REGION Network 92
   RUNG wire#powerrail
      Contact( "Carrier_14_Status.8" )
      Coil( "EMS".Carrier[14].SDC_IN.CrashDetectStatus )
   END_RUNG
   // the same network as SCL:
   "EMS".Carrier[14].SDC_IN.CrashDetectStatus := "Carrier_14_Status.8";
END_REGION

REGION Network 93
   RUNG wire#powerrail
      Contact( "Carrier_14_Status.9" )
      Coil( "EMS".Carrier[14].SDC_IN.EncoderCommFault )
   END_RUNG
   // the same network as SCL:
   "EMS".Carrier[14].SDC_IN.EncoderCommFault := "Carrier_14_Status.9";
END_REGION

REGION Network 94
   RUNG wire#powerrail
      Contact( "Carrier_14_Status.10" )
      Coil( "EMS".Carrier[14].SDC_IN.DriveCommFault )
   END_RUNG
   // the same network as SCL:
   "EMS".Carrier[14].SDC_IN.DriveCommFault := "Carrier_14_Status.10";
END_REGION

REGION Network 95
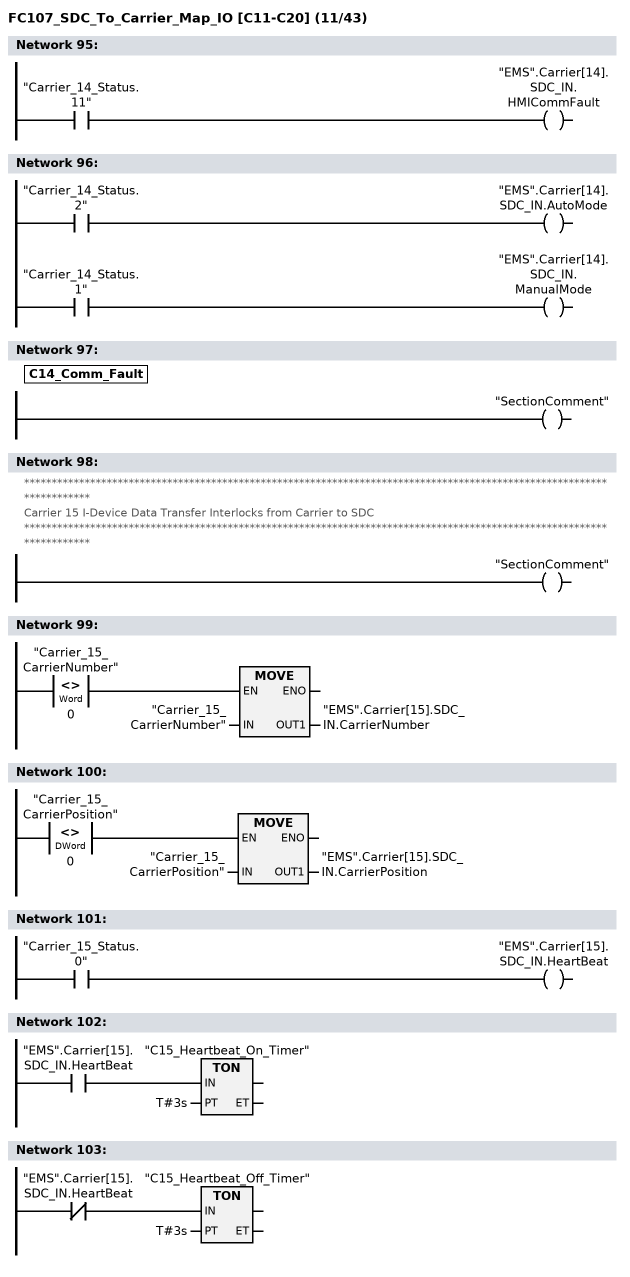
   RUNG wire#powerrail
      Contact( "Carrier_14_Status.11" )
      Coil( "EMS".Carrier[14].SDC_IN.HMICommFault )
   END_RUNG
   // the same network as SCL:
   "EMS".Carrier[14].SDC_IN.HMICommFault := "Carrier_14_Status.11";
END_REGION

REGION Network 96
   RUNG wire#powerrail
      Contact( "Carrier_14_Status.2" )
      Coil( "EMS".Carrier[14].SDC_IN.AutoMode )
   END_RUNG
   RUNG wire#powerrail
      Contact( "Carrier_14_Status.1" )
      Coil( "EMS".Carrier[14].SDC_IN.ManualMode )
   END_RUNG
   // the same network as SCL:
   "EMS".Carrier[14].SDC_IN.AutoMode := "Carrier_14_Status.2";
   "EMS".Carrier[14].SDC_IN.ManualMode := "Carrier_14_Status.1";
END_REGION

REGION Network 97
   Label( C14_Comm_Fault )
   RUNG wire#powerrail
      Coil( "SectionComment" )
   END_RUNG
   // the same network as SCL:
   C14_Comm_Fault:
   "SectionComment" := TRUE;
END_REGION

REGION Network 98
   // **********************************************************************************************************************
   // 
   // Carrier 15 I-Device Data Transfer Interlocks from Carrier to SDC
   // 
   // **********************************************************************************************************************
   RUNG wire#powerrail
      Coil( "SectionComment" )
   END_RUNG
   // the same network as SCL:
   "SectionComment" := TRUE;
END_REGION

REGION Network 99
   RUNG wire#powerrail
      { S7_Templates := "SrcType := Word" } NE_Contact(in1 := "Carrier_15_CarrierNumber", in2 := 0)
      Move(in := "Carrier_15_CarrierNumber", out1 => "EMS".Carrier[15].SDC_IN.CarrierNumber)
   END_RUNG
   // the same network as SCL:
   IF "Carrier_15_CarrierNumber" <> 0 THEN
       "EMS".Carrier[15].SDC_IN.CarrierNumber := "Carrier_15_CarrierNumber";
   END_IF;
END_REGION

REGION Network 100
   RUNG wire#powerrail
      { S7_Templates := "SrcType := DWord" } NE_Contact(in1 := "Carrier_15_CarrierPosition", in2 := 0)
      Move(in := "Carrier_15_CarrierPosition", out1 => "EMS".Carrier[15].SDC_IN.CarrierPosition)
   END_RUNG
   // the same network as SCL:
   IF "Carrier_15_CarrierPosition" <> 0 THEN
       "EMS".Carrier[15].SDC_IN.CarrierPosition := "Carrier_15_CarrierPosition";
   END_IF;
END_REGION

REGION Network 101
   RUNG wire#powerrail
      Contact( "Carrier_15_Status.0" )
      Coil( "EMS".Carrier[15].SDC_IN.HeartBeat )
   END_RUNG
   // the same network as SCL:
   "EMS".Carrier[15].SDC_IN.HeartBeat := "Carrier_15_Status.0";
END_REGION

REGION Network 102
   "C15_Heartbeat_On_Timer".TON(IN := "EMS".Carrier[15].SDC_IN.HeartBeat, PT := T#3s);
END_REGION

REGION Network 103
   "C15_Heartbeat_Off_Timer".TON(IN := NOT "EMS".Carrier[15].SDC_IN.HeartBeat, PT := T#3s);
END_REGION

REGION Network 104
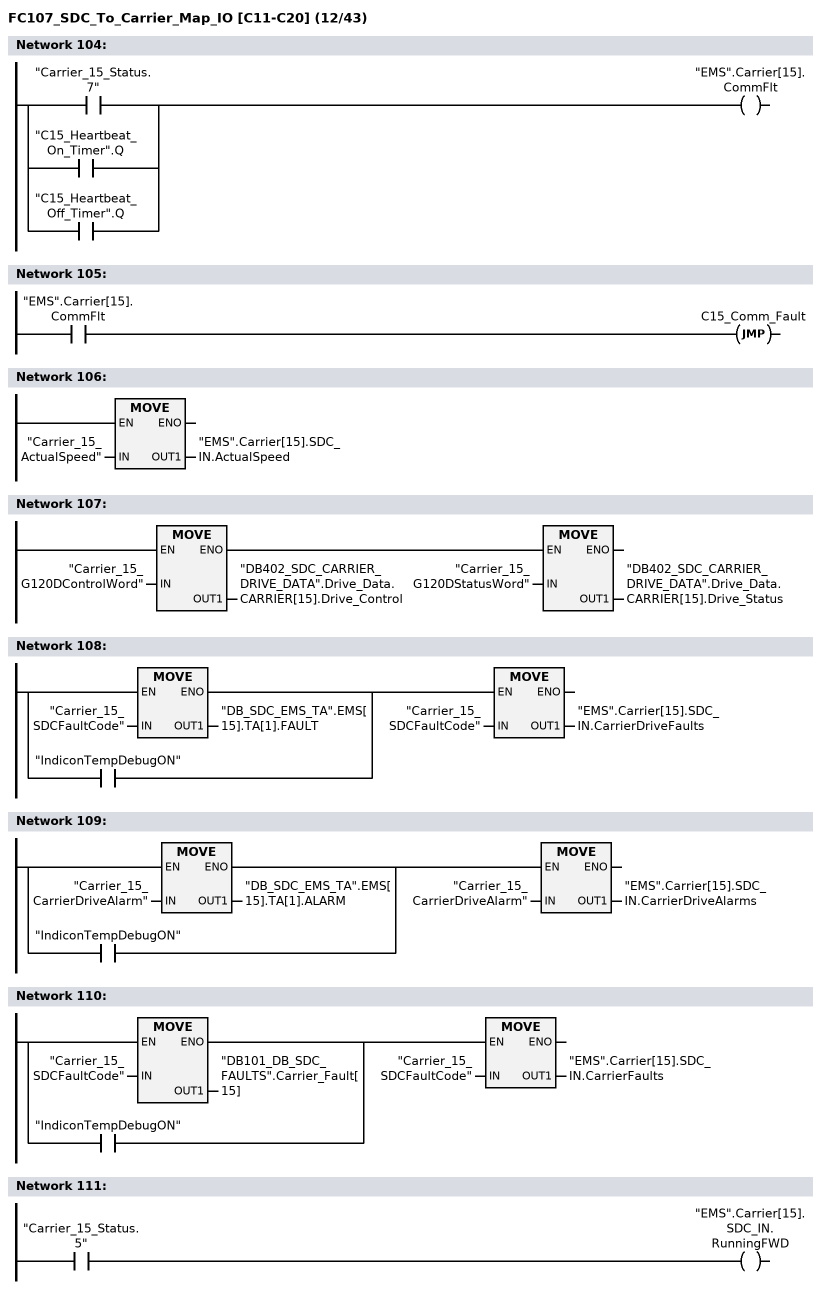
   RUNG wire#powerrail
      Contact( "Carrier_15_Status.7" )
      wire#w1
      Coil( "EMS".Carrier[15].CommFlt )
   END_RUNG
   RUNG wire#powerrail
      Contact( "C15_Heartbeat_On_Timer".Q )
   END_RUNG wire#w1
   RUNG wire#powerrail
      Contact( "C15_Heartbeat_Off_Timer".Q )
   END_RUNG wire#w1
   // the same network as SCL:
   "EMS".Carrier[15].CommFlt := "Carrier_15_Status.7" OR "C15_Heartbeat_On_Timer".Q OR "C15_Heartbeat_Off_Timer".Q;
END_REGION

REGION Network 105
   RUNG wire#powerrail
      Contact( "EMS".Carrier[15].CommFlt )
      JumpCoil( C15_Comm_Fault )
   END_RUNG
   // the same network as SCL:
   IF "EMS".Carrier[15].CommFlt THEN GOTO C15_Comm_Fault; END_IF;
END_REGION

REGION Network 106
   RUNG wire#powerrail
      Move(in := "Carrier_15_ActualSpeed", out1 => "EMS".Carrier[15].SDC_IN.ActualSpeed)
   END_RUNG
   // the same network as SCL:
   "EMS".Carrier[15].SDC_IN.ActualSpeed := "Carrier_15_ActualSpeed";
END_REGION

REGION Network 107
   RUNG wire#powerrail
      Move(in := "Carrier_15_G120DControlWord", out1 => "DB402_SDC_CARRIER_DRIVE_DATA".Drive_Data.CARRIER[15].Drive_Control)
      Move(in := "Carrier_15_G120DStatusWord", out1 => "DB402_SDC_CARRIER_DRIVE_DATA".Drive_Data.CARRIER[15].Drive_Status)
   END_RUNG
   // the same network as SCL:
   "DB402_SDC_CARRIER_DRIVE_DATA".Drive_Data.CARRIER[15].Drive_Control := "Carrier_15_G120DControlWord";
   "DB402_SDC_CARRIER_DRIVE_DATA".Drive_Data.CARRIER[15].Drive_Status := "Carrier_15_G120DStatusWord";
END_REGION

REGION Network 108
   RUNG wire#powerrail
      Move(in := "Carrier_15_SDCFaultCode", out1 => "DB_SDC_EMS_TA".EMS[15].TA[1].FAULT)
      wire#w1
      Move(in := "Carrier_15_SDCFaultCode", out1 => "EMS".Carrier[15].SDC_IN.CarrierDriveFaults)
   END_RUNG
   RUNG wire#powerrail
      Contact( "IndiconTempDebugON" )
   END_RUNG wire#w1
   // the same network as SCL:
   "DB_SDC_EMS_TA".EMS[15].TA[1].FAULT := "Carrier_15_SDCFaultCode";
   IF TRUE OR "IndiconTempDebugON" THEN
       "EMS".Carrier[15].SDC_IN.CarrierDriveFaults := "Carrier_15_SDCFaultCode";
   END_IF;
END_REGION

REGION Network 109
   RUNG wire#powerrail
      Move(in := "Carrier_15_CarrierDriveAlarm", out1 => "DB_SDC_EMS_TA".EMS[15].TA[1].ALARM)
      wire#w1
      Move(in := "Carrier_15_CarrierDriveAlarm", out1 => "EMS".Carrier[15].SDC_IN.CarrierDriveAlarms)
   END_RUNG
   RUNG wire#powerrail
      Contact( "IndiconTempDebugON" )
   END_RUNG wire#w1
   // the same network as SCL:
   "DB_SDC_EMS_TA".EMS[15].TA[1].ALARM := "Carrier_15_CarrierDriveAlarm";
   IF TRUE OR "IndiconTempDebugON" THEN
       "EMS".Carrier[15].SDC_IN.CarrierDriveAlarms := "Carrier_15_CarrierDriveAlarm";
   END_IF;
END_REGION

REGION Network 110
   RUNG wire#powerrail
      Move(in := "Carrier_15_SDCFaultCode", out1 => "DB101_DB_SDC_FAULTS".Carrier_Fault[15])
      wire#w1
      Move(in := "Carrier_15_SDCFaultCode", out1 => "EMS".Carrier[15].SDC_IN.CarrierFaults)
   END_RUNG
   RUNG wire#powerrail
      Contact( "IndiconTempDebugON" )
   END_RUNG wire#w1
   // the same network as SCL:
   "DB101_DB_SDC_FAULTS".Carrier_Fault[15] := "Carrier_15_SDCFaultCode";
   IF TRUE OR "IndiconTempDebugON" THEN
       "EMS".Carrier[15].SDC_IN.CarrierFaults := "Carrier_15_SDCFaultCode";
   END_IF;
END_REGION

REGION Network 111
   RUNG wire#powerrail
      Contact( "Carrier_15_Status.5" )
      Coil( "EMS".Carrier[15].SDC_IN.RunningFWD )
   END_RUNG
   // the same network as SCL:
   "EMS".Carrier[15].SDC_IN.RunningFWD := "Carrier_15_Status.5";
END_REGION

REGION Network 112
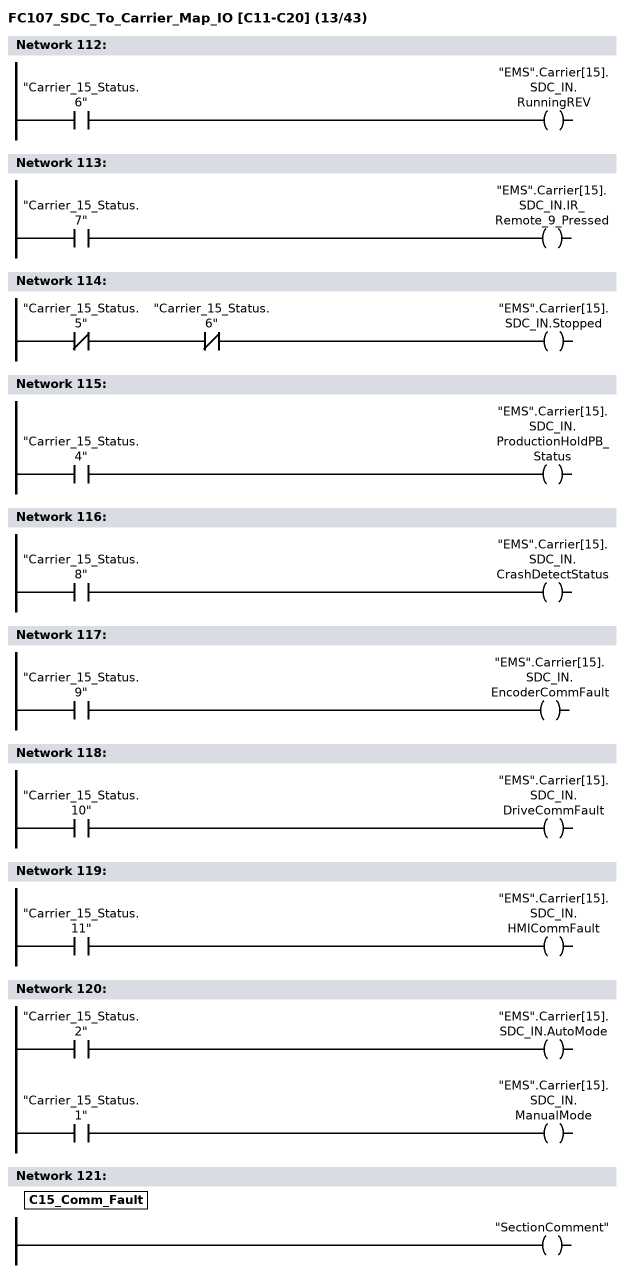
   RUNG wire#powerrail
      Contact( "Carrier_15_Status.6" )
      Coil( "EMS".Carrier[15].SDC_IN.RunningREV )
   END_RUNG
   // the same network as SCL:
   "EMS".Carrier[15].SDC_IN.RunningREV := "Carrier_15_Status.6";
END_REGION

REGION Network 113
   RUNG wire#powerrail
      Contact( "Carrier_15_Status.7" )
      Coil( "EMS".Carrier[15].SDC_IN.IR_Remote_9_Pressed )
   END_RUNG
   // the same network as SCL:
   "EMS".Carrier[15].SDC_IN.IR_Remote_9_Pressed := "Carrier_15_Status.7";
END_REGION

REGION Network 114
   RUNG wire#powerrail
      I_Contact( "Carrier_15_Status.5" )
      I_Contact( "Carrier_15_Status.6" )
      Coil( "EMS".Carrier[15].SDC_IN.Stopped )
   END_RUNG
   // the same network as SCL:
   "EMS".Carrier[15].SDC_IN.Stopped := NOT "Carrier_15_Status.5" AND NOT "Carrier_15_Status.6";
END_REGION

REGION Network 115
   RUNG wire#powerrail
      Contact( "Carrier_15_Status.4" )
      Coil( "EMS".Carrier[15].SDC_IN.ProductionHoldPB_Status )
   END_RUNG
   // the same network as SCL:
   "EMS".Carrier[15].SDC_IN.ProductionHoldPB_Status := "Carrier_15_Status.4";
END_REGION

REGION Network 116
   RUNG wire#powerrail
      Contact( "Carrier_15_Status.8" )
      Coil( "EMS".Carrier[15].SDC_IN.CrashDetectStatus )
   END_RUNG
   // the same network as SCL:
   "EMS".Carrier[15].SDC_IN.CrashDetectStatus := "Carrier_15_Status.8";
END_REGION

REGION Network 117
   RUNG wire#powerrail
      Contact( "Carrier_15_Status.9" )
      Coil( "EMS".Carrier[15].SDC_IN.EncoderCommFault )
   END_RUNG
   // the same network as SCL:
   "EMS".Carrier[15].SDC_IN.EncoderCommFault := "Carrier_15_Status.9";
END_REGION

REGION Network 118
   RUNG wire#powerrail
      Contact( "Carrier_15_Status.10" )
      Coil( "EMS".Carrier[15].SDC_IN.DriveCommFault )
   END_RUNG
   // the same network as SCL:
   "EMS".Carrier[15].SDC_IN.DriveCommFault := "Carrier_15_Status.10";
END_REGION

REGION Network 119
   RUNG wire#powerrail
      Contact( "Carrier_15_Status.11" )
      Coil( "EMS".Carrier[15].SDC_IN.HMICommFault )
   END_RUNG
   // the same network as SCL:
   "EMS".Carrier[15].SDC_IN.HMICommFault := "Carrier_15_Status.11";
END_REGION

REGION Network 120
   RUNG wire#powerrail
      Contact( "Carrier_15_Status.2" )
      Coil( "EMS".Carrier[15].SDC_IN.AutoMode )
   END_RUNG
   RUNG wire#powerrail
      Contact( "Carrier_15_Status.1" )
      Coil( "EMS".Carrier[15].SDC_IN.ManualMode )
   END_RUNG
   // the same network as SCL:
   "EMS".Carrier[15].SDC_IN.AutoMode := "Carrier_15_Status.2";
   "EMS".Carrier[15].SDC_IN.ManualMode := "Carrier_15_Status.1";
END_REGION

REGION Network 121
   Label( C15_Comm_Fault )
   RUNG wire#powerrail
      Coil( "SectionComment" )
   END_RUNG
   // the same network as SCL:
   C15_Comm_Fault:
   "SectionComment" := TRUE;
END_REGION

REGION Network 122
   // **********************************************************************************************************************
   // 
   // Carrier 16 I-Device Data Transfer Interlocks from Carrier to SDC
   // 
   // **********************************************************************************************************************
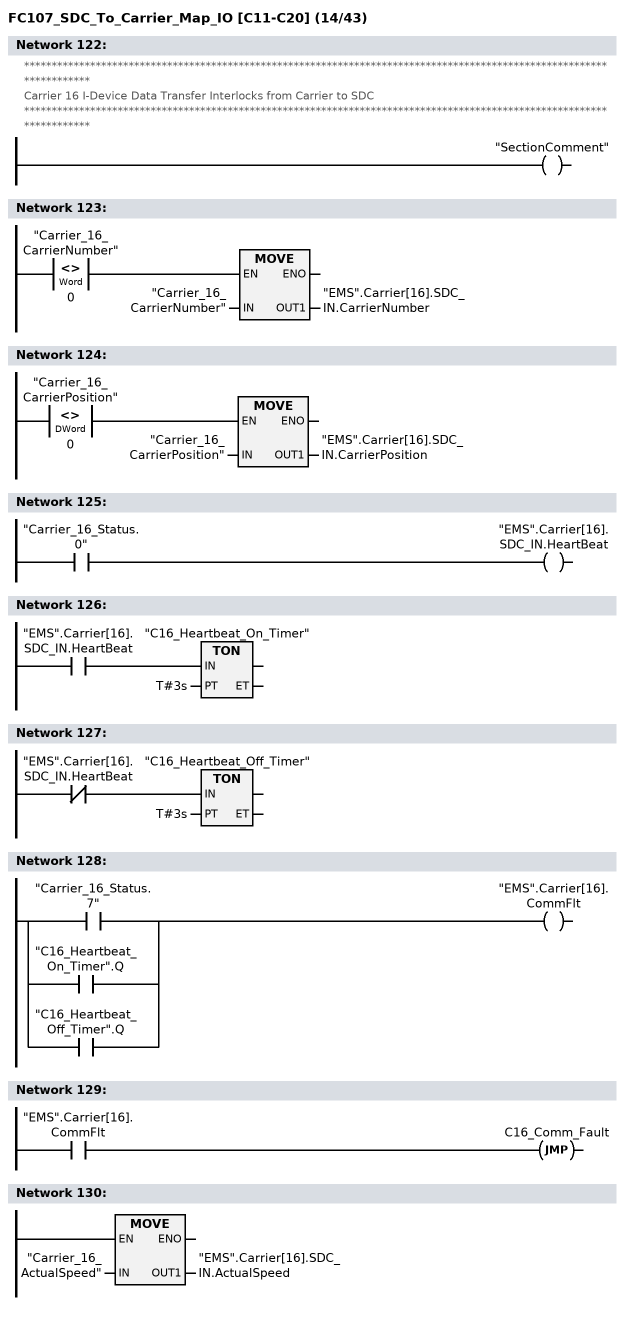
   RUNG wire#powerrail
      Coil( "SectionComment" )
   END_RUNG
   // the same network as SCL:
   "SectionComment" := TRUE;
END_REGION

REGION Network 123
   RUNG wire#powerrail
      { S7_Templates := "SrcType := Word" } NE_Contact(in1 := "Carrier_16_CarrierNumber", in2 := 0)
      Move(in := "Carrier_16_CarrierNumber", out1 => "EMS".Carrier[16].SDC_IN.CarrierNumber)
   END_RUNG
   // the same network as SCL:
   IF "Carrier_16_CarrierNumber" <> 0 THEN
       "EMS".Carrier[16].SDC_IN.CarrierNumber := "Carrier_16_CarrierNumber";
   END_IF;
END_REGION

REGION Network 124
   RUNG wire#powerrail
      { S7_Templates := "SrcType := DWord" } NE_Contact(in1 := "Carrier_16_CarrierPosition", in2 := 0)
      Move(in := "Carrier_16_CarrierPosition", out1 => "EMS".Carrier[16].SDC_IN.CarrierPosition)
   END_RUNG
   // the same network as SCL:
   IF "Carrier_16_CarrierPosition" <> 0 THEN
       "EMS".Carrier[16].SDC_IN.CarrierPosition := "Carrier_16_CarrierPosition";
   END_IF;
END_REGION

REGION Network 125
   RUNG wire#powerrail
      Contact( "Carrier_16_Status.0" )
      Coil( "EMS".Carrier[16].SDC_IN.HeartBeat )
   END_RUNG
   // the same network as SCL:
   "EMS".Carrier[16].SDC_IN.HeartBeat := "Carrier_16_Status.0";
END_REGION

REGION Network 126
   "C16_Heartbeat_On_Timer".TON(IN := "EMS".Carrier[16].SDC_IN.HeartBeat, PT := T#3s);
END_REGION

REGION Network 127
   "C16_Heartbeat_Off_Timer".TON(IN := NOT "EMS".Carrier[16].SDC_IN.HeartBeat, PT := T#3s);
END_REGION

REGION Network 128
   RUNG wire#powerrail
      Contact( "Carrier_16_Status.7" )
      wire#w1
      Coil( "EMS".Carrier[16].CommFlt )
   END_RUNG
   RUNG wire#powerrail
      Contact( "C16_Heartbeat_On_Timer".Q )
   END_RUNG wire#w1
   RUNG wire#powerrail
      Contact( "C16_Heartbeat_Off_Timer".Q )
   END_RUNG wire#w1
   // the same network as SCL:
   "EMS".Carrier[16].CommFlt := "Carrier_16_Status.7" OR "C16_Heartbeat_On_Timer".Q OR "C16_Heartbeat_Off_Timer".Q;
END_REGION

REGION Network 129
   RUNG wire#powerrail
      Contact( "EMS".Carrier[16].CommFlt )
      JumpCoil( C16_Comm_Fault )
   END_RUNG
   // the same network as SCL:
   IF "EMS".Carrier[16].CommFlt THEN GOTO C16_Comm_Fault; END_IF;
END_REGION

REGION Network 130
   RUNG wire#powerrail
      Move(in := "Carrier_16_ActualSpeed", out1 => "EMS".Carrier[16].SDC_IN.ActualSpeed)
   END_RUNG
   // the same network as SCL:
   "EMS".Carrier[16].SDC_IN.ActualSpeed := "Carrier_16_ActualSpeed";
END_REGION

REGION Network 131
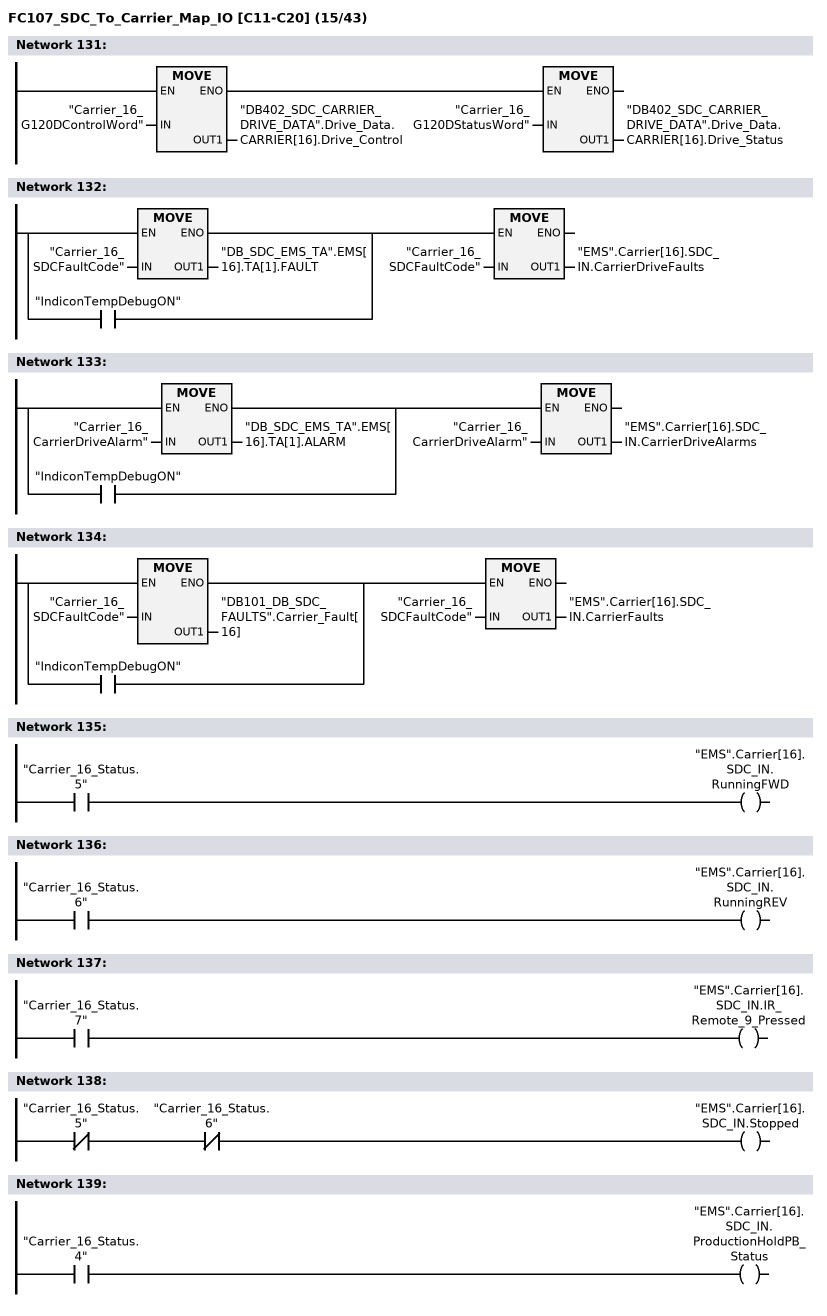
   RUNG wire#powerrail
      Move(in := "Carrier_16_G120DControlWord", out1 => "DB402_SDC_CARRIER_DRIVE_DATA".Drive_Data.CARRIER[16].Drive_Control)
      Move(in := "Carrier_16_G120DStatusWord", out1 => "DB402_SDC_CARRIER_DRIVE_DATA".Drive_Data.CARRIER[16].Drive_Status)
   END_RUNG
   // the same network as SCL:
   "DB402_SDC_CARRIER_DRIVE_DATA".Drive_Data.CARRIER[16].Drive_Control := "Carrier_16_G120DControlWord";
   "DB402_SDC_CARRIER_DRIVE_DATA".Drive_Data.CARRIER[16].Drive_Status := "Carrier_16_G120DStatusWord";
END_REGION

REGION Network 132
   RUNG wire#powerrail
      Move(in := "Carrier_16_SDCFaultCode", out1 => "DB_SDC_EMS_TA".EMS[16].TA[1].FAULT)
      wire#w1
      Move(in := "Carrier_16_SDCFaultCode", out1 => "EMS".Carrier[16].SDC_IN.CarrierDriveFaults)
   END_RUNG
   RUNG wire#powerrail
      Contact( "IndiconTempDebugON" )
   END_RUNG wire#w1
   // the same network as SCL:
   "DB_SDC_EMS_TA".EMS[16].TA[1].FAULT := "Carrier_16_SDCFaultCode";
   IF TRUE OR "IndiconTempDebugON" THEN
       "EMS".Carrier[16].SDC_IN.CarrierDriveFaults := "Carrier_16_SDCFaultCode";
   END_IF;
END_REGION

REGION Network 133
   RUNG wire#powerrail
      Move(in := "Carrier_16_CarrierDriveAlarm", out1 => "DB_SDC_EMS_TA".EMS[16].TA[1].ALARM)
      wire#w1
      Move(in := "Carrier_16_CarrierDriveAlarm", out1 => "EMS".Carrier[16].SDC_IN.CarrierDriveAlarms)
   END_RUNG
   RUNG wire#powerrail
      Contact( "IndiconTempDebugON" )
   END_RUNG wire#w1
   // the same network as SCL:
   "DB_SDC_EMS_TA".EMS[16].TA[1].ALARM := "Carrier_16_CarrierDriveAlarm";
   IF TRUE OR "IndiconTempDebugON" THEN
       "EMS".Carrier[16].SDC_IN.CarrierDriveAlarms := "Carrier_16_CarrierDriveAlarm";
   END_IF;
END_REGION

REGION Network 134
   RUNG wire#powerrail
      Move(in := "Carrier_16_SDCFaultCode", out1 => "DB101_DB_SDC_FAULTS".Carrier_Fault[16])
      wire#w1
      Move(in := "Carrier_16_SDCFaultCode", out1 => "EMS".Carrier[16].SDC_IN.CarrierFaults)
   END_RUNG
   RUNG wire#powerrail
      Contact( "IndiconTempDebugON" )
   END_RUNG wire#w1
   // the same network as SCL:
   "DB101_DB_SDC_FAULTS".Carrier_Fault[16] := "Carrier_16_SDCFaultCode";
   IF TRUE OR "IndiconTempDebugON" THEN
       "EMS".Carrier[16].SDC_IN.CarrierFaults := "Carrier_16_SDCFaultCode";
   END_IF;
END_REGION

REGION Network 135
   RUNG wire#powerrail
      Contact( "Carrier_16_Status.5" )
      Coil( "EMS".Carrier[16].SDC_IN.RunningFWD )
   END_RUNG
   // the same network as SCL:
   "EMS".Carrier[16].SDC_IN.RunningFWD := "Carrier_16_Status.5";
END_REGION

REGION Network 136
   RUNG wire#powerrail
      Contact( "Carrier_16_Status.6" )
      Coil( "EMS".Carrier[16].SDC_IN.RunningREV )
   END_RUNG
   // the same network as SCL:
   "EMS".Carrier[16].SDC_IN.RunningREV := "Carrier_16_Status.6";
END_REGION

REGION Network 137
   RUNG wire#powerrail
      Contact( "Carrier_16_Status.7" )
      Coil( "EMS".Carrier[16].SDC_IN.IR_Remote_9_Pressed )
   END_RUNG
   // the same network as SCL:
   "EMS".Carrier[16].SDC_IN.IR_Remote_9_Pressed := "Carrier_16_Status.7";
END_REGION

REGION Network 138
   RUNG wire#powerrail
      I_Contact( "Carrier_16_Status.5" )
      I_Contact( "Carrier_16_Status.6" )
      Coil( "EMS".Carrier[16].SDC_IN.Stopped )
   END_RUNG
   // the same network as SCL:
   "EMS".Carrier[16].SDC_IN.Stopped := NOT "Carrier_16_Status.5" AND NOT "Carrier_16_Status.6";
END_REGION

REGION Network 139
   RUNG wire#powerrail
      Contact( "Carrier_16_Status.4" )
      Coil( "EMS".Carrier[16].SDC_IN.ProductionHoldPB_Status )
   END_RUNG
   // the same network as SCL:
   "EMS".Carrier[16].SDC_IN.ProductionHoldPB_Status := "Carrier_16_Status.4";
END_REGION

REGION Network 140
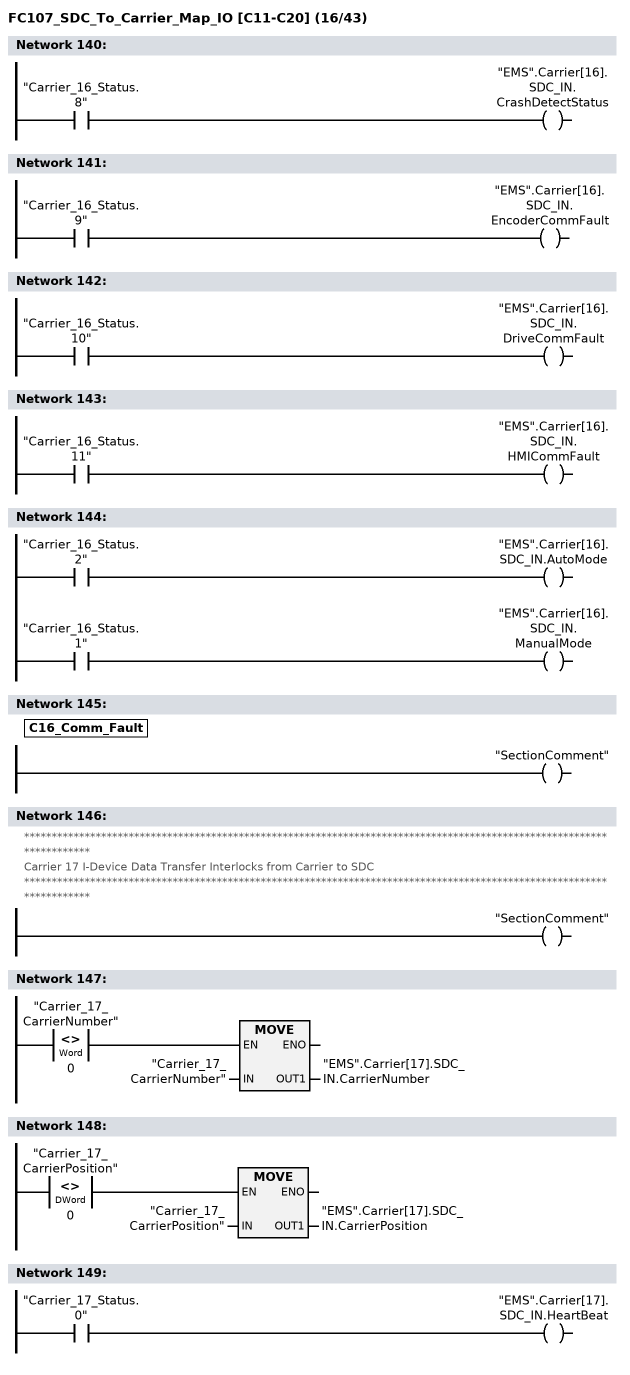
   RUNG wire#powerrail
      Contact( "Carrier_16_Status.8" )
      Coil( "EMS".Carrier[16].SDC_IN.CrashDetectStatus )
   END_RUNG
   // the same network as SCL:
   "EMS".Carrier[16].SDC_IN.CrashDetectStatus := "Carrier_16_Status.8";
END_REGION

REGION Network 141
   RUNG wire#powerrail
      Contact( "Carrier_16_Status.9" )
      Coil( "EMS".Carrier[16].SDC_IN.EncoderCommFault )
   END_RUNG
   // the same network as SCL:
   "EMS".Carrier[16].SDC_IN.EncoderCommFault := "Carrier_16_Status.9";
END_REGION

REGION Network 142
   RUNG wire#powerrail
      Contact( "Carrier_16_Status.10" )
      Coil( "EMS".Carrier[16].SDC_IN.DriveCommFault )
   END_RUNG
   // the same network as SCL:
   "EMS".Carrier[16].SDC_IN.DriveCommFault := "Carrier_16_Status.10";
END_REGION

REGION Network 143
   RUNG wire#powerrail
      Contact( "Carrier_16_Status.11" )
      Coil( "EMS".Carrier[16].SDC_IN.HMICommFault )
   END_RUNG
   // the same network as SCL:
   "EMS".Carrier[16].SDC_IN.HMICommFault := "Carrier_16_Status.11";
END_REGION

REGION Network 144
   RUNG wire#powerrail
      Contact( "Carrier_16_Status.2" )
      Coil( "EMS".Carrier[16].SDC_IN.AutoMode )
   END_RUNG
   RUNG wire#powerrail
      Contact( "Carrier_16_Status.1" )
      Coil( "EMS".Carrier[16].SDC_IN.ManualMode )
   END_RUNG
   // the same network as SCL:
   "EMS".Carrier[16].SDC_IN.AutoMode := "Carrier_16_Status.2";
   "EMS".Carrier[16].SDC_IN.ManualMode := "Carrier_16_Status.1";
END_REGION

REGION Network 145
   Label( C16_Comm_Fault )
   RUNG wire#powerrail
      Coil( "SectionComment" )
   END_RUNG
   // the same network as SCL:
   C16_Comm_Fault:
   "SectionComment" := TRUE;
END_REGION

REGION Network 146
   // **********************************************************************************************************************
   // 
   // Carrier 17 I-Device Data Transfer Interlocks from Carrier to SDC
   // 
   // **********************************************************************************************************************
   RUNG wire#powerrail
      Coil( "SectionComment" )
   END_RUNG
   // the same network as SCL:
   "SectionComment" := TRUE;
END_REGION

REGION Network 147
   RUNG wire#powerrail
      { S7_Templates := "SrcType := Word" } NE_Contact(in1 := "Carrier_17_CarrierNumber", in2 := 0)
      Move(in := "Carrier_17_CarrierNumber", out1 => "EMS".Carrier[17].SDC_IN.CarrierNumber)
   END_RUNG
   // the same network as SCL:
   IF "Carrier_17_CarrierNumber" <> 0 THEN
       "EMS".Carrier[17].SDC_IN.CarrierNumber := "Carrier_17_CarrierNumber";
   END_IF;
END_REGION

REGION Network 148
   RUNG wire#powerrail
      { S7_Templates := "SrcType := DWord" } NE_Contact(in1 := "Carrier_17_CarrierPosition", in2 := 0)
      Move(in := "Carrier_17_CarrierPosition", out1 => "EMS".Carrier[17].SDC_IN.CarrierPosition)
   END_RUNG
   // the same network as SCL:
   IF "Carrier_17_CarrierPosition" <> 0 THEN
       "EMS".Carrier[17].SDC_IN.CarrierPosition := "Carrier_17_CarrierPosition";
   END_IF;
END_REGION

REGION Network 149
   RUNG wire#powerrail
      Contact( "Carrier_17_Status.0" )
      Coil( "EMS".Carrier[17].SDC_IN.HeartBeat )
   END_RUNG
   // the same network as SCL:
   "EMS".Carrier[17].SDC_IN.HeartBeat := "Carrier_17_Status.0";
END_REGION

REGION Network 150
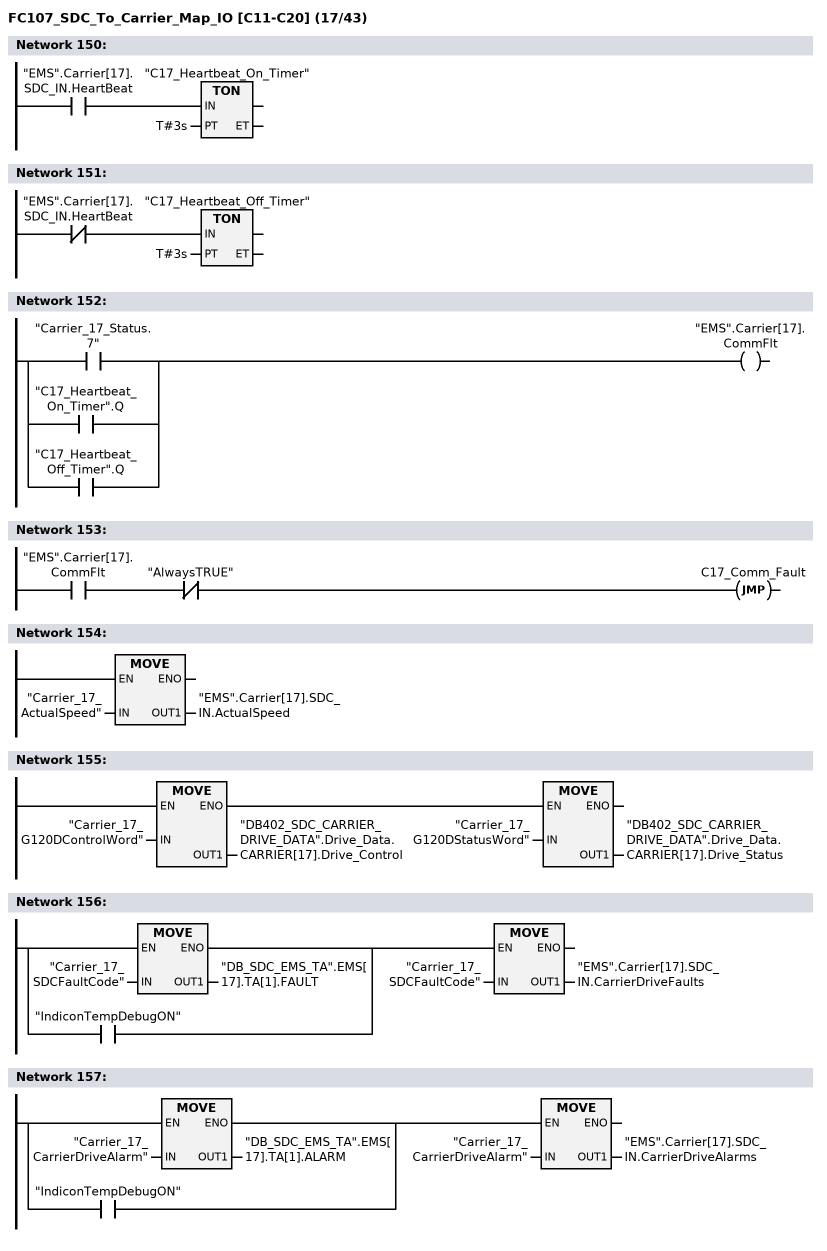
   "C17_Heartbeat_On_Timer".TON(IN := "EMS".Carrier[17].SDC_IN.HeartBeat, PT := T#3s);
END_REGION

REGION Network 151
   "C17_Heartbeat_Off_Timer".TON(IN := NOT "EMS".Carrier[17].SDC_IN.HeartBeat, PT := T#3s);
END_REGION

REGION Network 152
   RUNG wire#powerrail
      Contact( "Carrier_17_Status.7" )
      wire#w1
      Coil( "EMS".Carrier[17].CommFlt )
   END_RUNG
   RUNG wire#powerrail
      Contact( "C17_Heartbeat_On_Timer".Q )
   END_RUNG wire#w1
   RUNG wire#powerrail
      Contact( "C17_Heartbeat_Off_Timer".Q )
   END_RUNG wire#w1
   // the same network as SCL:
   "EMS".Carrier[17].CommFlt := "Carrier_17_Status.7" OR "C17_Heartbeat_On_Timer".Q OR "C17_Heartbeat_Off_Timer".Q;
END_REGION

REGION Network 153
   RUNG wire#powerrail
      Contact( "EMS".Carrier[17].CommFlt )
      I_Contact( "AlwaysTRUE" )
      JumpCoil( C17_Comm_Fault )
   END_RUNG
   // the same network as SCL:
   IF "EMS".Carrier[17].CommFlt AND NOT "AlwaysTRUE" THEN GOTO C17_Comm_Fault; END_IF;
END_REGION

REGION Network 154
   RUNG wire#powerrail
      Move(in := "Carrier_17_ActualSpeed", out1 => "EMS".Carrier[17].SDC_IN.ActualSpeed)
   END_RUNG
   // the same network as SCL:
   "EMS".Carrier[17].SDC_IN.ActualSpeed := "Carrier_17_ActualSpeed";
END_REGION

REGION Network 155
   RUNG wire#powerrail
      Move(in := "Carrier_17_G120DControlWord", out1 => "DB402_SDC_CARRIER_DRIVE_DATA".Drive_Data.CARRIER[17].Drive_Control)
      Move(in := "Carrier_17_G120DStatusWord", out1 => "DB402_SDC_CARRIER_DRIVE_DATA".Drive_Data.CARRIER[17].Drive_Status)
   END_RUNG
   // the same network as SCL:
   "DB402_SDC_CARRIER_DRIVE_DATA".Drive_Data.CARRIER[17].Drive_Control := "Carrier_17_G120DControlWord";
   "DB402_SDC_CARRIER_DRIVE_DATA".Drive_Data.CARRIER[17].Drive_Status := "Carrier_17_G120DStatusWord";
END_REGION

REGION Network 156
   RUNG wire#powerrail
      Move(in := "Carrier_17_SDCFaultCode", out1 => "DB_SDC_EMS_TA".EMS[17].TA[1].FAULT)
      wire#w1
      Move(in := "Carrier_17_SDCFaultCode", out1 => "EMS".Carrier[17].SDC_IN.CarrierDriveFaults)
   END_RUNG
   RUNG wire#powerrail
      Contact( "IndiconTempDebugON" )
   END_RUNG wire#w1
   // the same network as SCL:
   "DB_SDC_EMS_TA".EMS[17].TA[1].FAULT := "Carrier_17_SDCFaultCode";
   IF TRUE OR "IndiconTempDebugON" THEN
       "EMS".Carrier[17].SDC_IN.CarrierDriveFaults := "Carrier_17_SDCFaultCode";
   END_IF;
END_REGION

REGION Network 157
   RUNG wire#powerrail
      Move(in := "Carrier_17_CarrierDriveAlarm", out1 => "DB_SDC_EMS_TA".EMS[17].TA[1].ALARM)
      wire#w1
      Move(in := "Carrier_17_CarrierDriveAlarm", out1 => "EMS".Carrier[17].SDC_IN.CarrierDriveAlarms)
   END_RUNG
   RUNG wire#powerrail
      Contact( "IndiconTempDebugON" )
   END_RUNG wire#w1
   // the same network as SCL:
   "DB_SDC_EMS_TA".EMS[17].TA[1].ALARM := "Carrier_17_CarrierDriveAlarm";
   IF TRUE OR "IndiconTempDebugON" THEN
       "EMS".Carrier[17].SDC_IN.CarrierDriveAlarms := "Carrier_17_CarrierDriveAlarm";
   END_IF;
END_REGION

REGION Network 158
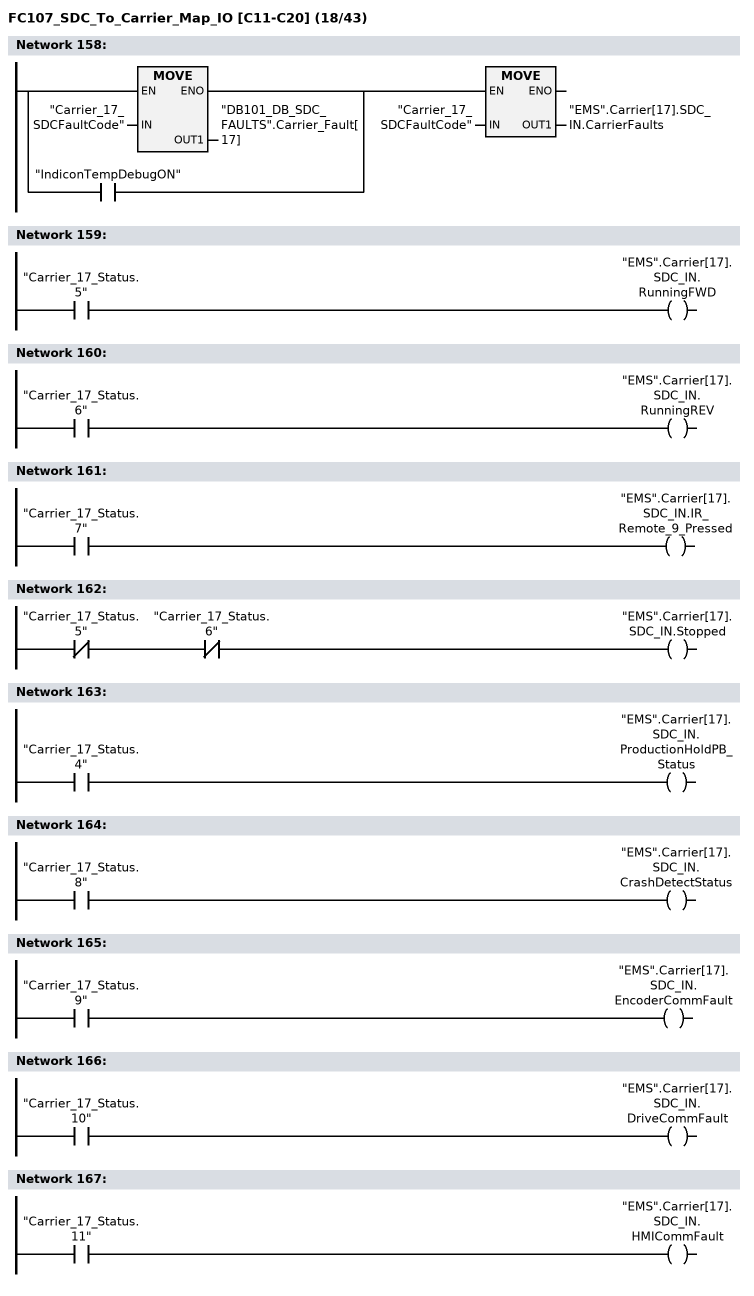
   RUNG wire#powerrail
      Move(in := "Carrier_17_SDCFaultCode", out1 => "DB101_DB_SDC_FAULTS".Carrier_Fault[17])
      wire#w1
      Move(in := "Carrier_17_SDCFaultCode", out1 => "EMS".Carrier[17].SDC_IN.CarrierFaults)
   END_RUNG
   RUNG wire#powerrail
      Contact( "IndiconTempDebugON" )
   END_RUNG wire#w1
   // the same network as SCL:
   "DB101_DB_SDC_FAULTS".Carrier_Fault[17] := "Carrier_17_SDCFaultCode";
   IF TRUE OR "IndiconTempDebugON" THEN
       "EMS".Carrier[17].SDC_IN.CarrierFaults := "Carrier_17_SDCFaultCode";
   END_IF;
END_REGION

REGION Network 159
   RUNG wire#powerrail
      Contact( "Carrier_17_Status.5" )
      Coil( "EMS".Carrier[17].SDC_IN.RunningFWD )
   END_RUNG
   // the same network as SCL:
   "EMS".Carrier[17].SDC_IN.RunningFWD := "Carrier_17_Status.5";
END_REGION

REGION Network 160
   RUNG wire#powerrail
      Contact( "Carrier_17_Status.6" )
      Coil( "EMS".Carrier[17].SDC_IN.RunningREV )
   END_RUNG
   // the same network as SCL:
   "EMS".Carrier[17].SDC_IN.RunningREV := "Carrier_17_Status.6";
END_REGION

REGION Network 161
   RUNG wire#powerrail
      Contact( "Carrier_17_Status.7" )
      Coil( "EMS".Carrier[17].SDC_IN.IR_Remote_9_Pressed )
   END_RUNG
   // the same network as SCL:
   "EMS".Carrier[17].SDC_IN.IR_Remote_9_Pressed := "Carrier_17_Status.7";
END_REGION

REGION Network 162
   RUNG wire#powerrail
      I_Contact( "Carrier_17_Status.5" )
      I_Contact( "Carrier_17_Status.6" )
      Coil( "EMS".Carrier[17].SDC_IN.Stopped )
   END_RUNG
   // the same network as SCL:
   "EMS".Carrier[17].SDC_IN.Stopped := NOT "Carrier_17_Status.5" AND NOT "Carrier_17_Status.6";
END_REGION

REGION Network 163
   RUNG wire#powerrail
      Contact( "Carrier_17_Status.4" )
      Coil( "EMS".Carrier[17].SDC_IN.ProductionHoldPB_Status )
   END_RUNG
   // the same network as SCL:
   "EMS".Carrier[17].SDC_IN.ProductionHoldPB_Status := "Carrier_17_Status.4";
END_REGION

REGION Network 164
   RUNG wire#powerrail
      Contact( "Carrier_17_Status.8" )
      Coil( "EMS".Carrier[17].SDC_IN.CrashDetectStatus )
   END_RUNG
   // the same network as SCL:
   "EMS".Carrier[17].SDC_IN.CrashDetectStatus := "Carrier_17_Status.8";
END_REGION

REGION Network 165
   RUNG wire#powerrail
      Contact( "Carrier_17_Status.9" )
      Coil( "EMS".Carrier[17].SDC_IN.EncoderCommFault )
   END_RUNG
   // the same network as SCL:
   "EMS".Carrier[17].SDC_IN.EncoderCommFault := "Carrier_17_Status.9";
END_REGION

REGION Network 166
   RUNG wire#powerrail
      Contact( "Carrier_17_Status.10" )
      Coil( "EMS".Carrier[17].SDC_IN.DriveCommFault )
   END_RUNG
   // the same network as SCL:
   "EMS".Carrier[17].SDC_IN.DriveCommFault := "Carrier_17_Status.10";
END_REGION

REGION Network 167
   RUNG wire#powerrail
      Contact( "Carrier_17_Status.11" )
      Coil( "EMS".Carrier[17].SDC_IN.HMICommFault )
   END_RUNG
   // the same network as SCL:
   "EMS".Carrier[17].SDC_IN.HMICommFault := "Carrier_17_Status.11";
END_REGION